// TIA Portal project "oscat_basic_332_s7_TIA_V12_V13_SP1_V14_V15.1" (V15.1) (continued)
VERSION : 1.1
// GEN_PW2 generates a time TH? followed by a time TL?.
// the input ts selects between 2 sets of timings for the operation.
// 
// uses: T_PLC_MS [FC64]
//       STIME [FB64],IDB_STIME [DB64]
   VAR_INPUT
      ENQ : Bool;
      TH1 : Time;
      TL1 : Time;
      TH2 : Time;
      TL2 : Time;
      TS : Bool;
   END_VAR
   VAR_OUTPUT
      Q : Bool;
      TH : Time;
      TL : Time;
   END_VAR
   VAR
      t_high : Time;
      t_low : Time;
      tx : Time;
      start : Time;
      init : Bool;
      et : Time;
   END_VAR
BEGIN


   (* read system timer *)
   #tx := T_CONV(DWORD_TO_DINT("T_PLC_MS"()));

   (* startup initialization *)
   IF NOT #init THEN
       #start := #tx;
       #init := TRUE;
       #TH := T#0s;
       #TL := T#0s;
   END_IF;

   (* timing selection *)
   IF #TS THEN
       #t_high := #TH2;
       #t_low := #TL2;
   ELSE
       #t_high := #TH1;
       #t_low := #TL1;
   END_IF;

   (* normal operation *)
   IF #ENQ THEN
       #et := #tx - #start;
       IF NOT #Q THEN
           IF #et >= #t_low THEN
               #Q := TRUE;
               #start := #tx;
               #TL := T#0s;
           ELSE
               #TL := #et;
           END_IF;
       ELSE
           IF #et >= #t_high THEN
               #Q := FALSE;
               #start := #tx;
               #TH := T#0s;
           ELSE
               #TH := #et;
           END_IF;
       END_IF;
   ELSE
       #Q := FALSE;
       #TH := T#0s;
       #TL := T#0s;
       #start := #tx;
   END_IF;


   (* revision history
   hm  26. sep. 2008   rev 1.0
       original version

   hm  14. mar. 2009   rev 1.1
       removed double assignments

   *)
END_FUNCTION_BLOCK

FUNCTION_BLOCK "GEN_RDM"   // FB97, SCL
TITLE = GEN_RDM
{ S7_Optimized_Access := 'FALSE' }
AUTHOR : oscat
FAMILY : SIGGEN
NAME : GEN_RDM
VERSION : 1.1
// this signal generator generates a random output. The signal is defined by period time (PT), 
// amplitude (AM), offset (OS).
// The Output waveform will have its max peak at AM/2 + OS and its minimum peak at -AM/2 + OS. 
// The period time PT defines how often the output signal will jump to a new randow value.
// The Output Q will be true for one cycle anytime the output OUT has changed
// 
// uses: T_PLC_MS [FC64]
//       STIME [FB64],IDB_STIME [DB64]
//       RDM [FC101]
//       BIT_COUNT [FC291] 
//       FRACT [FC83]
   VAR_INPUT
      PT : Time;
      AM : Real := 1.0e+0;
      OS : Real;
   END_VAR
   VAR_OUTPUT
      Q : Bool;
      Out : Real;
   END_VAR
   VAR
      tx : Time;
      last : Time;
      init : Bool;
   END_VAR
BEGIN


     (* read system time and prepare input data *)
     #tx := T_CONV(DWORD_TO_DINT("T_PLC_MS"())) - #last;

     (* init section *)
     IF NOT #init THEN
       #init := TRUE;
       #last := #tx;
       #tx := t#0s;
     END_IF;

     (* add last if one cycle is finished *)
     IF #tx >= #PT THEN
       #last := #last + #PT;
       #tx := #tx - #PT;

       (* generate output signal *)
       #Out := #AM * ("RDM"(0.0) - 0.5) + #OS;
       #Q := TRUE;
     ELSE
       #Q := FALSE;
     END_IF;

   (* revision history

   hm  7.2.2007    rev 1.0
     original version

   hm  16.9.2007    rev 1.1
     changes time() to T_plc_ms() for compatibility reasons

   *)
END_FUNCTION_BLOCK

FUNCTION_BLOCK "GEN_RDT"   // FB98, SCL
TITLE = GEN_RDT
{ S7_Optimized_Access := 'FALSE' }
AUTHOR : Schohaus
FAMILY : SIGGEN
NAME : GEN_RDT
VERSION : 1.1
// RDMT generates a defined pulse with pulse width TP_Q at random times. the random time will be defined with an minimum and maximum time.
// 
// uses: RDM [FC101]
//       T_PLC_MS [FC64] 
//       STIME [FB64],IDB_STIME [DB64] 
//       BIT_COUNT [FC291] 
//       FRACT [FC83]
   VAR_INPUT
      Enable : Bool := TRUE;
      Min_Time_ms : Time := T#1S;
      Max_Time_ms : Time := T#1S200MS;
      TP_Q : Time := T#100MS;
   END_VAR
   VAR_OUTPUT
      xQ : Bool;
   END_VAR
   VAR
      tonRDMTimer : TON;
      tof_xQ : TOF;
      tRDMTime : Time;
      rRDMTime : Real;
   END_VAR
BEGIN


   (*
   FUNCTION_BLOCK RDMTimer
   ###############################################################################
        Ersteller / author :                    J.Schohaus
        Datum / date:                         13.07.2007
   ###############################################################################
        Änderungen / Datum / Ersteller :                                                            
        moditication / date / author :        
   ###############################################################################
        Verwendete Bibliotheken     ( * werden im Baustein nicht benötigt )
                    Oscat.lib
   ###############################################################################
   Beschreibung:
   *)

     #tonRDMTimer ( IN:= #Enable , PT:= #tRDMTime );
     #tof_xQ ( IN:= #tonRDMTimer.Q , PT:= #TP_Q );
     #xQ := #tof_xQ.Q;
     IF #tonRDMTimer.Q THEN
          #xQ := TRUE ;
          #rRDMTime := "RDM" ( last:= #rRDMTime ) ;
          #tRDMTime := T_CONV(REAL_TO_DINT(#rRDMTime * DINT_TO_REAL(T_CONV(#Max_Time_ms - #Min_Time_ms)) + DINT_TO_REAL(T_CONV(#Min_Time_ms )))) ;
          #tonRDMTimer. IN:= FALSE ;
     END_IF;

   (* revision history
   J. Schohaus 19. nov 2007    rev 1.0
       origial version

   hm  16. mar. 2008           rev 1.1
       added type conversion to avoid warnings under codesys 3.0
   *)
END_FUNCTION_BLOCK

FUNCTION_BLOCK "GEN_RMP"   // FB99, SCL
TITLE = GEN_RMP
{ S7_Optimized_Access := 'FALSE' }
AUTHOR : oscat
FAMILY : SIGGEN
NAME : GEN_RMP
VERSION : 1.4
// this signal generator generates a ramp wave output. The ramp wave signal is defined by period time (PT), 
// amplitude (AM), offset (OS) and a specific delay for the output signal (DL).
// The Output waveform will have its minimum peak at OS and its maximum peak at AM + OS. 
// The delay input can delay a signal up to PT, this can be useful to synchronize different generators 
// and generate interleaving signals.
// in addition to the analog output Out there is a second boolean output Q with is true for one cycle when the ramp starts.
// 
// uses: T_PLC_MS [FC64]
//       STIME [FB64],IDB_STIME [DB64]
//       MODR [FC97]
//       FLOOR2 [FC82] 
//       FRACT [FC83]
//       MULTIME [FC203]
   VAR_INPUT
      PT : Time := T#1S;
      AM : Real := 1.0e+0;
      OS : Real;
      DL : Real;
   END_VAR
   VAR_OUTPUT
      Q : Bool;
      OUT : Real;
   END_VAR
   VAR
      tx : Time;
      last : Time;
      init : Bool;
      temp : Real;
      ltemp : Real;
   END_VAR
BEGIN


   (* read system time and prepare input data *)
   #tx := T_CONV(DWORD_TO_DINT("T_PLC_MS"())) - #last;
   #DL := "MODR"(IN:=#DL,DIVI:=1.0);
   IF #DL < 0.0 THEN #DL := 1.0 - #DL; END_IF;

   (* init section *)
   IF NOT #init THEN
       #init := TRUE;
       #last := #tx;
       #tx := t#0s;
   END_IF;

   (* add last if one cycle is finished *)
   IF #tx >= #PT THEN
       #last := #last + #PT;
       #tx := #tx - #PT;
   END_IF;

   (* generate sine wave *)
   #ltemp := #temp;
   IF #PT > t#0s THEN #temp := "FRACT"(DINT_TO_REAL(T_CONV(#tx + "MULTIME"(t:=#PT,M:=#DL))) / DINT_TO_REAL(T_CONV(#PT))); END_IF;
   #OUT := #AM * #temp + #OS;

   (* boolean output Q *)
   #Q := #temp < #ltemp;


   (* revision history
   hm  3. mar 2007     rev 1.0
       original version

   hm  17 sep 2007     rev 1.1
       replaced time() with t_plc_ms for compatibilitx reasons

   hm  27. nov 2007    rev 1.2
       avoid divide by 0 when pt = 0

   ks  26. oct. 2008   rev 1.3
       code optimization

   hm  10. mar. 2009   rev 1.4
       changed real constants to use dot syntax
   *)
END_FUNCTION_BLOCK

FUNCTION_BLOCK "GEN_SIN"   // FB100, SCL
TITLE = GEN_SIN
{ S7_Optimized_Access := 'FALSE' }
AUTHOR : oscat
FAMILY : SIGGEN
NAME : GEN_SIN
VERSION : 1.6
// this signal generator generates a sine wave output. The sine wave signal is defined by period time (PT), 
// amplitude (AM), offset (OS) and a specific delay for the output signal (DL).
// The Output waveform will have its max peak at AM/2 + OS and its minimum peak at -AM/2 + OS. 
// The delay input can delay a signal up to PT, this can be useful to synchronize different generators 
// and generate interleaving signals. A Cos wave can be generated accordingly.
// in addition to a analog output Out there is a second boolean output Q with the corresponding binary signal.
//  
// uses: T_PLC_MS [FC64]
//       STIME [FB64],IDB_STIME [DB64]
//       MODR [FC97]
//       FLOOR2 [FC82] 
//       MULTIME [FC203]
//       SIGN_R [FC109]
   VAR_INPUT
      PT : Time;
      AM : Real := 1.0e+0;
      OS : Real;
      DL : Real;
   END_VAR
   VAR_OUTPUT
      Q : Bool;
      OUT : Real;
   END_VAR
   VAR
      tx : Time;
      last : Time;
      init : Bool;
      temp : Real;
   END_VAR
BEGIN


   (* read system time and prepare input data *)
   #tx := T_CONV(DWORD_TO_DINT("T_PLC_MS"())) - #last;
   #DL := "MODR"(IN:=#DL,DIVI:=1.0);
   IF #DL < 0.0 THEN #DL := 1.0 - #DL; END_IF;

   (* init section *)
   IF NOT #init THEN
       #init := TRUE;
       #last := #tx;
       #tx := t#0s;
   END_IF;

   (* add last if one cycle is finished *)
   IF #tx >= #PT THEN
       #last := #last + #PT;
       #tx := #tx - #PT;
   END_IF;

   (* generate sine wave *)
   IF #PT > t#0s THEN #temp := SIN("PI2" * DINT_TO_REAL(T_CONV(#tx + "MULTIME"(t:=#PT,M:=#DL))) / DINT_TO_REAL(T_CONV(#PT))); END_IF;
   #OUT := #AM * 0.5 *  #temp + #OS;

   (* boolean output Q *)
   #Q := NOT "SIGN_R"(#temp);


   (* revision history
   hm  22. jan 2007    rev 1.0
       original version

   hm  17 sep 2007 rev 1.1
       replaced time() with t_plc_ms for compatibilitx reasons

   hm  27. nov 2007    rev 1.2
       avoid divide by 0 when pt = 0

   hm  6. jan 2008     rev 1.3
       improved performance

   hm  16. mar. 2008   rev 1.4
       added type conversion to avoid warnings under codesys 3.0

   hm  18. oct. 2008   rev 1.5
       using math constants

   hm  11. mar. 2009   rev 1.6
       changed real constants to use dot syntax

   *)
END_FUNCTION_BLOCK

FUNCTION_BLOCK "GEN_SQR"   // FB101, SCL
TITLE = GEN_SQR
{ S7_Optimized_Access := 'FALSE' }
AUTHOR : oscat
FAMILY : SIGGEN
NAME : GEN_SQR
VERSION : 1.4
// this signal generator generates a square wave output. The square wave signal is defined by period time (PT), 
// amplitude (AM), offset (OS), duty cycle (DC) and a specific delay for the output signal (DL).
// The Output waveform will switch between AM/2 + OS and -AM/2 + OS. The DC input specifies ther duty cycle, 
// DC = 0 means output is low at all times and 1 means output is high at all times.
// The delay input can delay a signal up to PT, this can be useful to synchronize different generators and generate interleaving signals.
// in addition to a analog output Out there is a second boolean output Q.
// 
// uses: T_PLC_MS [FC64]
//       STIME [FB64],IDB_STIME [DB64]
//       MODR [FC97]
//       FLOOR2 [FC82] 
//       MULTIME [FC203]
   VAR_INPUT
      PT : Time;
      AM : Real := 1.0e+0;
      OS : Real;
      DC : Real := 5.0e-1;
      DL : Real;
   END_VAR
   VAR_OUTPUT
      Q : Bool;
      Out : Real;
   END_VAR
   VAR
      tx : Time;
      last : Time;
      init : Bool;
   END_VAR
BEGIN


   (* check dc = 1 or 0 *)
   IF #DC = 0.0 THEN
       #Out := -#AM * 0.5 + #OS;
       #Q := FALSE;
       RETURN;
   ELSIF #DC = 1.0 THEN
       #Out := #AM * 0.5 + #OS;
       #Q := TRUE;
       RETURN;
   END_IF;

   (* read system time and prepare input data *)
   #tx := T_CONV(DWORD_TO_DINT("T_PLC_MS"())) - #last;
   #DL := "MODR"(IN:=#DL,DIVI:=1.0);
   IF #DL < 0.0 THEN #DL := 1.0 - #DL; END_IF;
   #DC := "MODR"(IN:=#DC,DIVI:=1.0);
   IF #DC < 0.0 THEN #DC := 1.0 - #DC; END_IF;

   (* init section *)
   IF NOT #init THEN
       #init := TRUE;
       #last := #tx;
       #tx := t#0s;
   END_IF;

   (* add last if one cycle is finished *)
   IF #tx >= #PT THEN
       #last := #last + #PT;
       #tx := #tx - #PT;
   END_IF;

   (* check if falling or rising edge first *)
   IF "MULTIME"(t:=#PT,M:=#DL + #DC) >= #PT THEN
       (* generate falling edge *)
       IF #tx >= "MULTIME"(t:=#PT,M:=#DL + #DC - 1) THEN
           #Out := -#AM * 0.5 + #OS;
           #Q := FALSE;
       END_IF;
       (* generate rising edge *)
       IF #tx >= "MULTIME"(t:=#PT,M:=#DL) THEN
           #Out := #AM * 0.5 + #OS;
           #Q := TRUE;
       END_IF;
   ELSE
       (* generate rising edge first *)
       IF #tx >= "MULTIME"(t:=#PT,M:=#DL) THEN
           #Out := #AM * 0.5 + #OS;
           #Q := TRUE;
       END_IF;
       (* generate falling edge *)
       IF #tx >= "MULTIME"(t:=#PT,M:=#DL + #DC) THEN
           #Out := -#AM * 0.5 + #OS;
           #Q := FALSE;
       END_IF;
   END_IF;


   (* revision history

   hm  12. feb 2007    rev 1.1
       added default value for dc = 0.5

   hm  17 sep 2007 rev 1.2
       replaced time() with t_plc_ms for compatibilitx reasons

   hm  6. jan 2008 rev 1.3
       improved performance

   hm  11. mar. 2009   rev 1.4
       changed real constants to use dot syntax
       set default amplitude to 1.0

   *)
END_FUNCTION_BLOCK

FUNCTION_BLOCK "PWM_DC"   // FB102, SCL
TITLE = PWM_DC
{ S7_Optimized_Access := 'FALSE' }
AUTHOR : oscat
FAMILY : SIGGEN
NAME : PWM_DC
VERSION : 1.4
// this signal generator generates a square wave signal which is specified by the frequency and the duty cycle
// 
// uses: CLK_PRG [FB52]
//       T_PLC_MS [FC64] 
//       STIME [FB64],IDB_STIME [DB64] 
//       TP_X [FB69]
   VAR_INPUT
      F : Real;
      DC : Real;
   END_VAR
   VAR_OUTPUT
      Q : Bool;
   END_VAR
   VAR
      clk : "CLK_PRG";
      pulse : "TP_X";
   END_VAR
   VAR_TEMP
      tmp : Real;
   END_VAR
BEGIN


   IF #F > 0.0 THEN
       #tmp := 1000.0 / #F;
       #clk(PT := T_CONV(REAL_TO_DINT(#tmp)));
       #pulse(IN := #clk.Q, PT := T_CONV(REAL_TO_DINT(#tmp * #DC)));
       #Q := #pulse.Q;
   END_IF;


   (* revision history

   hm  25. feb 2007    rev 1.1
       recoded in st for better performance and better portability

   hm  27. nov 2007    rev 1.2
       avoid divide by 0 when F = 0

   hm  19. oct. 2008   rev 1.3
       changed type TP_R to TP_X because of name change
       improved performance

   hm  11. mar. 2009   rev 1.4
       changed real constants to use dot syntax

   *)
END_FUNCTION_BLOCK

FUNCTION_BLOCK "PWM_PW"   // FB103, SCL
TITLE = PWM_PW
{ S7_Optimized_Access := 'FALSE' }
AUTHOR : oscat
FAMILY : SIGGEN
NAME : PWM_PW
VERSION : 1.5
// this signal generator generates a square wave signal which is specified by the frequency and the pulse width.
// 
// uses: CLK_PRG [FB52]
//       T_PLC_MS [FC64] 
//       STIME [FB64],IDB_STIME [DB64] 
//       TP_X [FB69]
   VAR_INPUT
      F : Real;
      PW : Time;
   END_VAR
   VAR_OUTPUT
      Q : Bool;
   END_VAR
   VAR
      clk : "CLK_PRG";
      pulse : "TP_X";
   END_VAR
BEGIN


   IF #F > 0.0 THEN
       #clk(PT := T_CONV(REAL_TO_DINT(1000.0 / #F)));
       #pulse(IN := #clk.Q, PT := #PW);
       #Q := #pulse.Q;
   END_IF;


   (* revision history

   hm  25. feb 2007    rev 1.1
       recoded in st for better performance and better portability

   hm  27. nov 2007    rev 1.2
       avoid divide by 0 when F = 0

   hm  9. dec 2007     rev 1.3
       corrected an error with F = 0

   hm  19. oct. 2008   rev 1.4
       changed type tp_r to TP_x brecause of name change

   hm  11. mar. 2009   rev 1.5
       changed real constants to use dot syntax

   *)
END_FUNCTION_BLOCK

FUNCTION_BLOCK "RMP_SOFT"   // FB104, SCL
TITLE = RMP_SOFT
{ S7_Optimized_Access := 'FALSE' }
AUTHOR : oscat
FAMILY : SIGGEN
NAME : RMP_SOFT
VERSION : 2.0
// this soft on/off ramp generator generates a soft on and soft off ramp while the max on value is set by the input
// the time for a full ramp can be set by config variables for up and down ramp.
// 
// uses: _RMP_B [FB93]
//       T_PLC_MS [FC64] 
//       STIME [FB64],IDB_STIME [DB64]
   VAR_INPUT
      IN : Bool;
      VAL : Byte;
      PT_ON : Time;
      PT_OFF : Time;
   END_VAR
   VAR_OUTPUT
      OUT : Byte;
   END_VAR
   VAR
      rmp : "_RMP_B";
      tmp : Byte;
   END_VAR
BEGIN


   #tmp := INT_TO_BYTE(SEL(G:=#IN, IN0:=0, IN1:=BYTE_TO_INT(#VAL)));
   IF BYTE_TO_INT(#tmp) > BYTE_TO_INT(#OUT) THEN
       (* we need to ramp down *)
       #rmp(DIR := TRUE, E := TRUE, TR := #PT_ON, RMP := #OUT);
       (* make sure out does not surpass tmp *)
       #OUT := INT_TO_BYTE(MIN(IN1:=BYTE_TO_INT(#OUT), IN2:=BYTE_TO_INT(#tmp)));
   ELSIF BYTE_TO_INT(#tmp) < BYTE_TO_INT(#OUT) THEN
       (* we need to ramp up *)
       #rmp(DIR := FALSE, E := TRUE, TR := #PT_OFF, RMP := #OUT);
       (* make sure out does not surpass tmp *)
       #OUT := INT_TO_BYTE(MAX(IN1:=BYTE_TO_INT(#OUT), IN2:=BYTE_TO_INT(#tmp)));
   ELSE
       (* no ramp necessary *)
       #rmp(E := FALSE, RMP := #OUT);
   END_IF;


   (* revision history

   hm 22.1.2007    rev 1.1
       deleted unused variables X1 and I, X2 and X3

   hm  17.9.2007   rev 1.2
       replaced time() with t_plc_ms() for compatibility reasons

   hm  26. oct. 2008   2.0
       new code using _rmp_b
   *)
END_FUNCTION_BLOCK

FUNCTION_BLOCK "RMP_W"   // FB105, SCL
TITLE = RMP_W
{ S7_Optimized_Access := 'FALSE' }
AUTHOR : oscat
FAMILY : SIGGEN
NAME : RMP_W
VERSION : 2.0
// this ramp generator generates a Word wide ramp with 65535 steps
// the generator has an asynchronous set and reset
// the ramp is controlled by PT which is the total ramp time for a full sweep from 0..65535
// an UD input controlls the direction Up or Down and the E input enables the ramp generation
// a busy output indicates that the ramp is running, busy false means output is stable.
// the outputs low and high will be true when the output has reached its max or min value.
// 
// uses: _RMP_W [FB94]
//       T_PLC_MS [FC64] 
//       STIME [FB64],IDB_STIME [DB64]
   VAR_INPUT
      SET : Bool;
      PT : Time;
      "E" : Bool := TRUE;
      UP : Bool := TRUE;
      RST : Bool;
   END_VAR
   VAR_OUTPUT
      out : Word;
      busy : Bool;
      high : Bool;
      low : Bool;
   END_VAR
   VAR
      rmp : "_RMP_W";
   END_VAR
BEGIN


   #rmp(DIR := #UP, E := #"E", TR := #PT, RMP := #out);

   (* set or reset operation *)
   IF #RST THEN
       #out := 0;
   ELSIF #SET THEN
       #out := 65535;
   END_IF;

   (* checks for outputs stable and reset or set busy flag *)
   #low := #out = 0;
   #high := #out = 65535;
   #busy := NOT (#low OR #high) AND #"E";


   (* revision history:

   hm 4.10.2006        rev 1.1
       added the busy output which signals that the ramp is running.

   hm 22.1.2007        rev 1.2
       deleted unused variable step

   hm  17.9.2007       rev 1.3
       replaced time() with t_plc_ms() for compatibility reasons

   hm  28. sep 2007    rev 1.4
       added outputs on and off
       busy is now disabled while en is false
       new coding for higher accuracy and performance

   hm  5. oct 2007 rev 1.5
       added statements to allow for PT to be t#0s output jumps to max or min immediately

   hm  2. dec 2007 rev 1.6
       corrected an error in calculation of step response

   hm  25. dec 2007    rev 1.7
       corrected an error while step response was too slow for fast rise times

   hm  16. oct. 2008   rev 1.8
       improved performance

   hm  18. oct. 2008   rev 1.9
       renamed inout EN to E for compatibility reasons

   hm  23. oct. 2008   rev 2.0
       new code using _RMP_W
   *)
END_FUNCTION_BLOCK

FUNCTION_BLOCK "RMP_B"   // FB232, SCL
TITLE = RMP_B
{ S7_Optimized_Access := 'FALSE' }
AUTHOR : oscat
FAMILY : SIGGEN
NAME : RMP_B
VERSION : 2.0
// this ramp generator generates a byte wide ramp with 255 steps
// the generator has an asynchronous set and reset
// the ramp is controlled by PT which is the total ramp time for a full sweep from 0..255
// an UD input controlls the direction Up or Down and the E input enables the ramp generation
// a busy output indicates that the ramp is running, busy false means output is stable.
// the outputs low and high will be true when the output has reached its max or min value.
// 
// uses: _RMP_B [FB93]
//       T_PLC_MS [FC64] 
//       STIME [FB64],IDB_STIME [DB64]
   VAR_INPUT
      SET : Bool;
      PT : Time;
      "E" : Bool := TRUE;
      UP : Bool := TRUE;
      RST : Bool;
   END_VAR
   VAR_OUTPUT
      OUT : Byte;
      BUSY : Bool;
      HIGH : Bool;
      LOW : Bool;
   END_VAR
   VAR
      rmp : "_RMP_B";
   END_VAR
BEGIN


   (* generate ramp *)
   #rmp(DIR := #UP, E := #"E", TR := #PT, RMP := #OUT);

   (* set or reset operation *)
   IF #RST THEN
       #OUT := 0;
   ELSIF #SET THEN
       #OUT := 255;
   END_IF;

   (* checks for outputs stable and reset or set busy flag *)
   #LOW := #OUT = 0;
   #HIGH := #OUT = 255;
   #BUSY := NOT (#LOW OR #HIGH) AND #"E";


   (* revision history

   hm 5.10.2006    rev 1.1
       added busy output
   hm 17.1.2007    rev 1.2
       renamed input ud to up for better usability
       deleted unused variable step

   hm  17.9.2007       rev 1.3
       replaced time() with t_plc_ms() for compatibility reasons

   hm  28. sep 2007    rev 1.4
       added outputs on and off
       busy is now disabled while en is false
       new coding for higher accuracy and performance

   hm  5. oct 2007 rev 1.5
       added statements to allow for PT to be t#0s output jumps to max or min immediately

   hm  25. dec 2007    rev 1.6
       improved code for better performance

   hm  16. oct. 2008   rev 1.7
       improved code for better performance

   hm  18. oct. 2008   rev 1.8
       added type conversion to avoid warnings
       changed input en to e for compatibility reasons

   hm  23. oct. 2008   REV     2.0
       new code using _RMP_B

   *)
END_FUNCTION_BLOCK

FUNCTION_BLOCK "TREND_DW"   // FB245, SCL
TITLE = TREND_DW
{ S7_Optimized_Access := 'FALSE' }
AUTHOR : hugo
FAMILY : SIGPRO
NAME : TREND_DW
VERSION : 1.2
// trend_DW analyses the trend of a input signal.
// The Output Q is True if the input X is >= last_X and is false if the input X is <= last_X
// in addition to the trend the output TU will be high for one cycle to signal a rising of the input value X
// and  TD will signal a decreasing value on the input X.
// in case of a change the output D will show the delta of the input to the last input value.
   VAR_INPUT
      X : DWord;
   END_VAR
   VAR_OUTPUT
      Q : Bool;
      TU : Bool;
      TD : Bool;
      D : DWord;
   END_VAR
   VAR
      last_X : DWord;
   END_VAR
BEGIN


   IF DWORD_TO_DINT(#X) > DWORD_TO_DINT(#last_X) THEN
       #TU := TRUE;
       #TD := FALSE;
       #D := DINT_TO_DWORD(DWORD_TO_DINT(#X) - DWORD_TO_DINT(#last_X));
       #Q := TRUE;
   ELSIF DWORD_TO_DINT(#X) < DWORD_TO_DINT(#last_X) THEN
       #TD := TRUE;
       #TU := FALSE;
       #D := DINT_TO_DWORD(DWORD_TO_DINT(#last_X) - DWORD_TO_DINT(#X));
       #Q := FALSE;
   ELSE
       #TU := FALSE; 
       #TD := FALSE;
       #D := 0;
   END_IF;
   #last_X := #X;


   (* revision history
   hm  21. nov. 2008   rev 1.0
       original version

   hm  20. feb. 2009   rev 1.1
       added outputs TU, TD and D

   hm  14. mar. 2009   rev 1.2
       removed double assignments

   *)
END_FUNCTION_BLOCK

FUNCTION_BLOCK "_RMP_NEXT"   // FB246, SCL
TITLE = _RMP_NEXT
{ S7_Optimized_Access := 'FALSE' }
AUTHOR : hugo
FAMILY : SIGGEN
NAME : RMP_NEXT
VERSION : 1.4
// _RMP_NEXT  will generate a ramp output following the input IN.
// on a rising ramp the output will stop as soon as it has surpassed the input in, and on a falling ramp it will stop when out is smaller than in.
// a lockout time T_L will be added between up and down direction.
// 
// uses: _RMP_B [FB93]
//       TREND_DW [FB245]
//       T_PLC_MS [FC64]
//       STIME [FB64],IDB_STIME [DB64]
   VAR_INPUT
      "E" : Bool := TRUE;
      IN : Byte;
      TR : Time;
      TF : Time;
      TL : Time;
   END_VAR
   VAR_OUTPUT
      DIR : Bool;
      UP : Bool;
      DN : Bool;
   END_VAR
   VAR_IN_OUT
      OUT : Byte;
   END_VAR
   VAR
      rmx : "_RMP_B";
      dirx : "TREND_DW";
      t_lock : TP;
      xen : Bool;
      xdir : Bool;
   END_VAR
BEGIN


   #dirx(X := #IN);

   #t_lock(IN := FALSE, PT := #TL);

   IF #dirx.TU AND (BYTE_TO_INT(#OUT) < BYTE_TO_INT(#IN)) THEN
       IF NOT #xdir AND #xen THEN #t_lock.IN := TRUE; END_IF;
       #xen := TRUE;
       #xdir := TRUE;
   ELSIF #dirx.TD AND (BYTE_TO_INT(#OUT) > BYTE_TO_INT(#IN)) THEN
       IF #xdir AND #xen THEN #t_lock.IN := TRUE; END_IF;
       #xen := TRUE;
       #xdir := FALSE;
   ELSIF #xen THEN
       IF (#xdir AND (BYTE_TO_INT(#OUT) >= BYTE_TO_INT(#IN))) OR (NOT #xdir AND (BYTE_TO_INT(#OUT) <= BYTE_TO_INT(#IN))) THEN
           #xen := FALSE;
           IF #TL > t#0s THEN #t_lock.IN := TRUE; END_IF;
       END_IF;
   END_IF;

   IF NOT #t_lock.Q AND #xen THEN
       #UP := #xdir; 
       #DIR := #xdir;
       #DN := NOT #xdir;
   ELSE
       #DN := FALSE;
       #UP := FALSE; 
   END_IF;

   #rmx(RMP := #OUT, E := #"E" AND (#UP OR #DN) , DIR := #DIR, TR := SEL(G:=#DIR, IN0:=#TF, IN1:=#TR));


   (* revison history
   hm  23. nov. 2008 rev 1.0
     original version

   hm  24. jan. 2009 rev 1.1
     deleted unused vars tmp1, tmp2

   hm  20. feb. 2009 rev 1.2
     improved algorithm
     added TL

   hm  9. mar. 2009  rev 1.3
     input E was ignored
     removed double assignments

   hm  18. jul. 2009 rev 1.4
     improved performance

   *)
END_FUNCTION_BLOCK

FUNCTION "T_PLC_MS" : DWord   // FC64, SCL
TITLE = T_PLC_MS
{ S7_Optimized_Access := 'FALSE' }
AUTHOR : hugo
FAMILY : MEASURE
NAME : T_PLC_MS
VERSION : 1.2
// T_PLC_MS reads the internal PLC timer and return the time, it has the advantage to be able to set a debug mode 
// and speed up the counter to test the plc timer overrun which occurs every 50 days respectively 25 days at siemens S7
// this routine also allows to correct the behavior of s7 where the internal plc counter will not count all 32 bits.
// 
// uses: STIME [FB64],IDB_STIME [DB64]
BEGIN


   "IDB_STIME"(); 
   #T_PLC_MS := "IDB_STIME".tx; 
   (* hier muss die korrektur für step7 stattfinden
   plctime muss den vollen wertebereich von time ausnutzen:
   wenn bei step7 time -24tage bis plus 24 tage ist dann muss der timer auch beim überlauf auf -24tage springen 
   und auf keinen fall auf 0 !!!!
   für siemens muss ein weiterer fb im main eingebunden werden der sicherstellt das alle 32 bits durchgezählt werden.
   es kann nur ein fb sein den er muss sich das oberste (32te) bit merken.
   oder etwa spring s7 bei überlauf auf -24 tage????? dann wäre keine korrektur nötig.
   *)
   IF "debug" THEN
       #T_PLC_MS := DINT_TO_DWORD((DWORD_TO_DINT(SHL(IN:=#T_PLC_MS,N:="N") OR SHL(IN:=DWORD#1,N:="N"))-1) + DWORD_TO_DINT("offset_1"));
   END_IF;


   (* revision history
   hm  14.9.2007   rev 1.0
       original version

   hm  12. nov 2007    rev 1.1
       added temporaray variable tx because some compilers could not handle time() as an argument

   hm  16. nov. 2008   rev 1.2
       initialized constants with 0 for compatibility reasons
   *)
END_FUNCTION

FUNCTION "FLOOR2" : DInt   // FC82, SCL
TITLE = FLOOR2
{ S7_Optimized_Access := 'FALSE' }
AUTHOR : hugo
FAMILY : MATH
NAME : FLOOR2
VERSION : 1.1
// This is a rounding function which returns the biggest possible integer which is less or equal to X.
// floor2(3.14) = 3
// floor2(-3.14) = -4
   VAR_INPUT
      X : Real;
   END_VAR
BEGIN


   #FLOOR2 := REAL_TO_DINT(#X);
   IF DINT_TO_REAL(#FLOOR2) > #X THEN
     #FLOOR2 := #FLOOR2 - 1;
   END_IF;

   (* revision history
   hm  21. mar. 2008   rev 1.0
       originlal version

   hm  4. apr. 2008    rev 1.1
       added type conversion to avoid warnings under codesys 3.0
   *)
END_FUNCTION

FUNCTION "FRACT" : Real   // FC83, SCL
TITLE = FRACT
{ S7_Optimized_Access := 'FALSE' }
AUTHOR : hugo
FAMILY : MATH
NAME : FRACT
VERSION : 1.3
// this function returns the fraction of a real number
// fract(3.14) = 0.14
   VAR_INPUT
      x : Real;
   END_VAR
BEGIN


   IF ABS(#x) < 2.0E9 THEN
       #FRACT := #x - DINT_TO_REAL(TRUNC(#x));
   ELSE
       #FRACT := 0.0;
   END_IF;


   (* revision history
   hm  4. aug 2006 rev 1.0
       original version

   hm  11. mar 2008    rev 1.1
       added dint_to_real for compatibility reasons
       now returns 0 for number > 2e9
       changed input to x

   hm  21. mar. 2008   rev 1.2
       use D_trunc instead of TRUNC for compatibility reasons

   hm  10. mar. 2009   rev 1.3
       real constants updated to new systax using dot

   *)
END_FUNCTION

FUNCTION "MODR" : Real   // FC97, SCL
TITLE = MODR
{ S7_Optimized_Access := 'FALSE' }
AUTHOR : hugo
FAMILY : MATH
NAME : MODR
VERSION : 1.5
// this is a modulo funtion for real numbers
// modr(5.5,2.5) = 0.5
// 
// uses: FLOOR2 [FC82]
   VAR_INPUT
      IN : Real;
      DIVI : Real;
   END_VAR
BEGIN


   IF #DIVI = 0.0 THEN
       #MODR := 0.0;
   ELSE
       #MODR := #IN - DINT_TO_REAL("FLOOR2"(#IN / #DIVI)) * #DIVI;
   END_IF;


   (* revision history

   hm  4. aug.2006     rev 1.0

   hm  28. jan.2007   rev 1.1
       modr(x,0) will deliver the result 0

   hm  21. mar 2008    rev 1.2
       use D_trunc for compatibility reasons

   hm  4. apr. 2008    rev 1.3
       added type conversion to avoid warnings under codesys 3.0

   hm  31. oct. 2008   rev 1.4
       changed algorithm to the more common version using floor instead of TRUNC

   hm  10. mar. 2009   rev 1.5
       real constants updated to new systax using dot

   *)
END_FUNCTION

FUNCTION "RDM" : Real   // FC101, SCL
TITLE = RDM
{ S7_Optimized_Access := 'FALSE' }
AUTHOR : hugo
FAMILY : MATH
NAME : RDM
VERSION : 1.9
// this function calculates a pseudo random number
// to generate the number it reads the sps timer and calculates a random number between 0 and 1:
// in order to use rdm more then once within one sps cycle it need to be called with different seed numbers LAST.
//  
// uses: T_PLC_MS [FC64]
//       STIME [FB64],IDB_STIME [DB64]
//       BIT_COUNT [FC291]
//       FRACT [FC83]
   VAR_INPUT
      last : Real;
   END_VAR
   VAR_TEMP
      tn : DWord;
      _tn AT tn : Array[0..31] of Bool;
      tc : Int;
   END_VAR
BEGIN


   #tn := "T_PLC_MS"();
   #tc := "BIT_COUNT"(#tn);
   #_tn[7] := #_tn[26];  //tn.31 := tn.2;
   #_tn[6] := #_tn[29];  //tn.30 := tn.5;
   #_tn[5] := #_tn[28];  //tn.29 := tn.4;
   #_tn[4] := #_tn[25];  //tn.28 := tn.1;
   #_tn[3] := #_tn[24];  //tn.27 := tn.0;
   #_tn[2] := #_tn[31];  //tn.26 := tn.7;
   #_tn[1] := #_tn[30];  //tn.25 := tn.6;
   #_tn[0] := #_tn[27];  //tn.24 := tn.3;
   #tn := ROL(IN:=#tn,N:="BIT_COUNT"(#tn)) AND 16#7FFFFFFF OR 16#40000001;  // OR 16#80000001
   #tn := DINT_TO_DWORD(DWORD_TO_DINT(#tn) MOD 71474513 + #tc + 77);
   #RDM := "FRACT"(DINT_TO_REAL(DWORD_TO_DINT(#tn)) / 10000000.0 * ("E"- LIMIT(MN:=0.0,IN:=#last,MX:=1.0)));


   (*
   pt := ADR(temp);
   pt^ := (T_PLC_MS() AND 16#007FFFFF) OR 16#3D000000;
   RDM := fract(modR(temp*e+pi1, PI1-last) + modR(temp*PI1+e + last,e-last));
   *)

   (* revision history
   hm      16. jan 2007        rev 1.0
       original version

   hm      11. nov 2007        rev 1.1
       changed time() into t_plc_ms()

   hm      20. nov 2007        rev 1.2
       changed code of temp calculation to avoid overflow in modr due to resuclt would not fit DINT for high timeer values

   hm      5. jan 2008     rev 1.3
       changed calculation of temp to avoid problem with high values of t_plc_ms

   hm      2. feb 2008     rev 1.4
       changed algorithm to avoind non iec functions and guarantee more randomness

   hm  10. mar. 2008       rev 1.5
       make sure last will be between 0 and 1 to avoid invalid results

   hm  16. mar. 2008       rev 1.6
       added conversion for tc to avoid warnings under codesys 3.0

   hm  18. may. 2008       rev 1.7
       changed constant E to E1

   hm  18. oct. 2008       rev 1.8
       using math constants

   hm  10. mar. 2009       rev 1.9
       real constants updated to new systax using dot

   *)
END_FUNCTION

FUNCTION "SIGN_R" : Bool   // FC109, SCL
TITLE = SIGN_R
{ S7_Optimized_Access := 'FALSE' }
AUTHOR : hugo
FAMILY : MATH
NAME : SIGN_R
VERSION : 1.4
// this function return true if the real input is negative
   VAR_INPUT
      in : Real;
   END_VAR
BEGIN


   #SIGN_R := #in < 0.0;


   (* revision history
   hm 19.1.2007    rev 1.1
       changed method of function for better compatibility to other systems

   hm  1.12.2007   rev 1.2
       changed code to improve performance

   hm  14. jun. 2008   rev 1.3
       improved performace

   hm 10. mar. 2009    rev 1.4
       real constants updated to new systax using dot
   *)
END_FUNCTION

FUNCTION "MULTIME" : Time   // FC203, SCL
TITLE = MULTIME
{ S7_Optimized_Access := 'FALSE' }
AUTHOR : hugo
FAMILY : TIDT
NAME : MULTIME
VERSION : 1.1
// multiplies a time by a real number and returns a time
   VAR_INPUT
      t : Time;
      "M" : Real;
   END_VAR
BEGIN


     #MULTIME := T_CONV(REAL_TO_DINT(DINT_TO_REAL(T_CONV(#t))*#"M"));

   (* revision history
   hm      2. oct 2006 rev 1.0
       original version

   hm      14. mar 2008    rev 1.1
       rounded the result after the last digit

   *)
END_FUNCTION

FUNCTION "BIT_COUNT" : Int   // FC291, SCL
TITLE = BIT_COUNT
{ S7_Optimized_Access := 'FALSE' }
AUTHOR : hugo
FAMILY : GATE
NAME : BITCT
VERSION : 1.1
// BIT_COUNT counts the amount True of bits in a dword.
// for exabple: bit_count(3) returns 2 because two bits (bits 0 and 1) are true and all others are false.
   VAR_INPUT
      IN : DWord;
   END_VAR
   VAR_TEMP
      temp : DWord;
      attemp AT temp : Array[0..31] of Bool;
   END_VAR
BEGIN


     #BIT_COUNT := 0;
     #temp := #IN;

     WHILE DWORD_TO_DINT(#temp) <> 0 DO
       IF #attemp[24] THEN #BIT_COUNT := #BIT_COUNT +1; END_IF;
       #temp := SHR(IN:=#temp,N:=1);
     END_WHILE;

   (* revision history
   5.7.2007  rev 1.0    original version

   10.9.2007  rev 1.1    hm
     changed algorithm for better performace
     the execution time has reduced by a factor of 5
     deleted unused variable temp
   *)
END_FUNCTION

FUNCTION "FRMP_B" : Byte   // FC424, SCL
TITLE = FRMP_B
{ S7_Optimized_Access := 'FALSE' }
AUTHOR : hugo
FAMILY : FUNCT
NAME : FRMP_B
VERSION : 1.0
// this function calculates a ramp and limits the output to 0 .. 255 without overflow problems
   VAR_INPUT
      START : Byte;
      DIR : Bool;
      TD : Time;
      TR : Time;
   END_VAR
   VAR_TEMP
      tTD : Time;
   END_VAR
BEGIN


   #tTD := #TD;  // only Step7

   IF #TD < #TR THEN
     #FRMP_B := DINT_TO_BYTE(MIN(IN1:=DWORD_TO_DINT(SHL(IN:=DINT_TO_DWORD(T_CONV(#tTD)), N:=8)) / T_CONV(#TR) 
                                ,IN2:=SEL(G:=#DIR, IN0:=BYTE_TO_DINT(#START), IN1:=BYTE_TO_DINT(BYTE#255) - BYTE_TO_DINT(#START))));
     IF #DIR THEN
       #FRMP_B := INT_TO_BYTE(BYTE_TO_INT(#START) + BYTE_TO_INT(#FRMP_B));
     ELSE
       #FRMP_B := INT_TO_BYTE(BYTE_TO_INT(#START) - BYTE_TO_INT(#FRMP_B));
     END_IF;
   ELSE
     #FRMP_B := INT_TO_BYTE(DINT_TO_INT(SEL(G:=#DIR, IN0:=0, IN1:=255)));
   END_IF;


   (* revision history

   17. feb. 2011 rev 1.0
     new module

   *)
END_FUNCTION

// ===== PLC "Eng signal processing"  Unspecific CPU S7 300 =====

VAR_GLOBAL CONSTANT   // PLC tag table "STEP7 classic symbols"
   "debug" : Bool := FALSE;
   "N" : Int := 0;
   "offset_FC64" : Int := 0;   // MigChange: offset
   "ff" : DWord := 16#FFFFFFFF;
   "ff_FC318" : Byte := 2#1;   // MigChange: ff
   "offset_FC64_1" : DWord := 0;
END_VAR

DATA_BLOCK "IDB_STIME"   // DB64
{ S7_Optimized_Access := 'FALSE' }
AUTHOR : dalbi
FAMILY : MEASURE
VERSION : 0.0
// stored: InstanceOfName STIME
"STIME"
BEGIN
END_DATA_BLOCK

FUNCTION_BLOCK "STIME"   // FB64, SCL
TITLE = STIME
{ S7_Optimized_Access := 'FALSE' }
AUTHOR : dalbi
FAMILY : MEASURE
NAME : STIME
VERSION : 1.5
// this function block makes sure that the timer of a siemens sps counts from 0 - 2^32-1.
   VAR_OUTPUT
      tx : DWord;
      at_tx AT tx : Array[0..31] of Bool;
   END_VAR
   VAR
      last_time : DWord;
      bit31 : Bool;
      init : Bool := TRUE;
   END_VAR
   VAR_TEMP
      TOP_SI : Struct
         EV_CLASS : Byte;
         EV_NUM : Byte;
         PRIORITY : Byte;
         NUM : Byte;
         TYP2_3 : Byte;
         TYP1 : Byte;
         ZI1 : Word;
         ZI2_3 : DWord;
      END_STRUCT;
      START_UP_SI : Struct
         EV_CLASS : Byte;
         EV_NUM : Byte;
         PRIORITY : Byte;
         NUM : Byte;
         TYP2_3 : Byte;
         TYP1 : Byte;
         ZI1 : Word;
         ZI2_3 : DWord;
      END_STRUCT;
      ERR : Int;
   END_VAR
BEGIN


   (* this FB is only necessary for siemens sps
   the siemens sps timer counts from 0 to 2^31-1 and starts at 0 sfter overrun.
   this means that the bit 31 (the highest bit ) will never be used and therefore
   a problem arises when t2 - t1 is checked.
   t2 - t1 is always valid also in an timer overrun situation where the time t1 is very high and t2 is very low.
   the result of the subtraction t2 - t1 however is still valid.
   this calculation does not work for soiemens because the highest bit is not used.

   this module stores the highest bit, changes the highest bit at every overrun occurence and stuffs ther highest bit in the output.
   the output is then used by t_plc_us and t_plc_ms.

   the correction needs and fb and not a function because the value of the highest bit has to be stored.

   do never use this function block in a codesys environment. the timer in codesys is correct and runs from 0 to 2^32-1
   *)

   (* read actual startup info *)
   (* OB1_SCAN_1  BYTE  -  B#16#01: Abschluss des Neustarts (Warmstarts)
                        -  B#16#02: Abschluss des Wiederanlaufs
                        -  B#16#03: Abschluss des freien Zyklus
                        -  B#16#04: Abschluss des Kaltstarts
                        -  B#16#05: Erster OB 1-Zyklus der neuen Master-CPU nach 
                                    Master-Reserve-Umschaltung und STOP des 
                                    bisherigen Masters *)

   #ERR := RD_SINFO (TOP_SI => #TOP_SI, START_UP_SI => #START_UP_SI);

   (* reset last_time on system startup *)
   IF #TOP_SI.EV_NUM = 1 OR #TOP_SI.EV_NUM = 2 OR #TOP_SI.EV_NUM = 4 OR NOT #init THEN 
       #last_time := 0;
       #bit31 := false;
       #init := true;
   END_IF;

   (* read the system timer *)
   #tx := DINT_TO_DWORD(T_CONV(TIME_TCK()));

   (* stuff the highest bit into the timer value *)
   #at_tx[7] := #bit31;

   (* check for overrun *)
   IF DWORD_TO_DINT(#tx) < DWORD_TO_DINT(#last_time) THEN
       (* an overrun has occured, change the value of the highest bit *)
       #bit31 := NOT #bit31;
   END_IF;

   (* stuff the highest bit into the timer value *)
   #at_tx[7] := #bit31;

   (* remember the last system time for the next overrun check *)
   #last_time := #tx;


   (* revision history
   DA  14.9.2007 rev 1.0
     original version

   DA  24.2.2008 rev 1.1
     added self reset on system startup

   DA   2.5.2008 rev 1.2
     correct a problem running under OB35

   DA  12.3.2009 rev 1.3
     correct a problem run on different CPUs

   DA  22.12.2009 rev 1.4
     correct a problem on startup

   DA  19.09.2011 rev 1.5
     correct a error in code 
   *)
END_FUNCTION_BLOCK

FUNCTION_BLOCK "_RMP_W"   // FB94, SCL
TITLE = _RMP_W
{ S7_Optimized_Access := 'FALSE' }
AUTHOR : hugo
FAMILY : SIGGEN
NAME : _RMP_W
VERSION : 1.1
// _RMP_B generates a ramp on an external var of type byte
// tr is the total ramp time, E is an enable and dir the direction of the ramp
// 
// uses: T_PLC_MS [FC64]
//       STIME [FB64],IDB_STIME [DB64]
   VAR_INPUT
      DIR : Bool;
      "E" : Bool := TRUE;
      TR : Time;
   END_VAR
   VAR_IN_OUT
      RMP : Word;
   END_VAR
   VAR
      tx : DWord;
      tl : DWord;
      "step" : DInt;
      init : Bool;
      last_dir : Bool;
   END_VAR
   VAR_TEMP
      TOP_SI : Struct
         EV_CLASS : Byte;
         EV_NUM : Byte;
         PRIORITY : Byte;
         NUM : Byte;
         TYP2_3 : Byte;
         TYP1 : Byte;
         ZI1 : Word;
         ZI2_3 : DWord;
      END_STRUCT;
      START_UP_SI : Struct
         EV_CLASS : Byte;
         EV_NUM : Byte;
         PRIORITY : Byte;
         NUM : Byte;
         TYP2_3 : Byte;
         TYP1 : Byte;
         ZI1 : Word;
         ZI2_3 : DWord;
      END_STRUCT;
      ERR : Int;
   END_VAR
BEGIN


   (* read actual startup info *)
   (* OB1_SCAN_1  BYTE  -  B#16#01: Abschluss des Neustarts (Warmstarts)
                        -  B#16#02: Abschluss des Wiederanlaufs
                        -  B#16#03: Abschluss des freien Zyklus
                        -  B#16#04: Abschluss des Kaltstarts
                        -  B#16#05: Erster OB 1-Zyklus der neuen Master-CPU nach 
                                    Master-Reserve-Umschaltung und STOP des 
                                    bisherigen Masters *)

   #ERR := RD_SINFO (TOP_SI => #TOP_SI, START_UP_SI => #START_UP_SI);

   (* reset last_time on system startup *)
   IF #TOP_SI.EV_NUM = 1 OR #TOP_SI.EV_NUM = 2 OR #TOP_SI.EV_NUM = 4 THEN 
       #init := FALSE;
   END_IF;

   #tx := "T_PLC_MS"();
   IF #"E" AND #init THEN
       (* we need to set tl = tx when direction changes *)
       IF #DIR XOR #last_dir THEN
        #tl := #tx;
        #last_dir := #DIR;
       END_IF;
       (* check_elapsed time and calculate only if necessary *)
       IF #TR > t#0s THEN
           #"step" := DWORD_TO_DINT(SHL(IN:=DINT_TO_DWORD(DWORD_TO_DINT(#tx)-DWORD_TO_DINT(#tl)), N:=16)) / T_CONV(#TR);
       ELSE
           #"step" := 65535;
       END_IF;
       IF #"step" > 0 THEN
           (* perform the step on the ramp *)
           #tl := #tx;
           (* calculate the step response *)
           IF NOT #DIR THEN #"step" := - #"step"; END_IF;
           #RMP := DINT_TO_WORD(LIMIT(MN:=0, IN:=WORD_TO_DINT(#RMP) + #"step", MX:=65535));
       END_IF;
   ELSE
       #tl := #tx;
       #init := TRUE;
   END_IF;


   (* revison history
   hm  22. oct. 2008   rev 1.0
       original version

   hm  20. nov. 2008   rev 1.1
       set default for E to be TRUE
       added init

   *)
END_FUNCTION_BLOCK

FUNCTION_BLOCK "RMP_W"   // FB105, SCL
TITLE = RMP_W
{ S7_Optimized_Access := 'FALSE' }
AUTHOR : oscat
FAMILY : SIGGEN
NAME : RMP_W
VERSION : 2.0
// this ramp generator generates a Word wide ramp with 65535 steps
// the generator has an asynchronous set and reset
// the ramp is controlled by PT which is the total ramp time for a full sweep from 0..65535
// an UD input controlls the direction Up or Down and the E input enables the ramp generation
// a busy output indicates that the ramp is running, busy false means output is stable.
// the outputs low and high will be true when the output has reached its max or min value.
// 
// uses: _RMP_W [FB94]
//       T_PLC_MS [FC64] 
//       STIME [FB64],IDB_STIME [DB64]
   VAR_INPUT
      SET : Bool;
      PT : Time;
      "E" : Bool := TRUE;
      UP : Bool := TRUE;
      RST : Bool;
   END_VAR
   VAR_OUTPUT
      out : Word;
      busy : Bool;
      high : Bool;
      low : Bool;
   END_VAR
   VAR
      rmp : "_RMP_W";
   END_VAR
BEGIN


   #rmp(DIR := #UP, E := #"E", TR := #PT, RMP := #out);

   (* set or reset operation *)
   IF #RST THEN
       #out := 0;
   ELSIF #SET THEN
       #out := 65535;
   END_IF;

   (* checks for outputs stable and reset or set busy flag *)
   #low := #out = 0;
   #high := #out = 65535;
   #busy := NOT (#low OR #high) AND #"E";


   (* revision history:

   hm 4.10.2006        rev 1.1
       added the busy output which signals that the ramp is running.

   hm 22.1.2007        rev 1.2
       deleted unused variable step

   hm  17.9.2007       rev 1.3
       replaced time() with t_plc_ms() for compatibility reasons

   hm  28. sep 2007    rev 1.4
       added outputs on and off
       busy is now disabled while en is false
       new coding for higher accuracy and performance

   hm  5. oct 2007 rev 1.5
       added statements to allow for PT to be t#0s output jumps to max or min immediately

   hm  2. dec 2007 rev 1.6
       corrected an error in calculation of step response

   hm  25. dec 2007    rev 1.7
       corrected an error while step response was too slow for fast rise times

   hm  16. oct. 2008   rev 1.8
       improved performance

   hm  18. oct. 2008   rev 1.9
       renamed inout EN to E for compatibility reasons

   hm  23. oct. 2008   rev 2.0
       new code using _RMP_W
   *)
END_FUNCTION_BLOCK

FUNCTION_BLOCK "AIN1"   // FB106, SCL
TITLE = AIN1
{ S7_Optimized_Access := 'FALSE' }
AUTHOR : oscat
FAMILY : SIGPRO
NAME : AIN1
VERSION : 1.3
// Ain1 converts signals from A/D converters or other digital sources to an internal real value.
   VAR_INPUT
      in : DWord;
      sign_bit : Int := 255;
      error_bit : Int := 255;
      error_code_EN : Bool;
      error_code : DWord;
      overflow_bit : Int := 255;
      overflow_code_en : Bool;
      overflow_code : DWord;
      Bit_0 : Int;
      Bit_N : Int := 31;
      out_min : Real;
      out_max : Real := 1.0e+1;
      code_min : DWord;
      code_max : DWord := DW#16#FFFFFFFF;
      error_output : Real;
      overflow_output : Real := 1.0e+1;
   END_VAR
   VAR_OUTPUT
      out : Real;
      sign : Bool;
      error : Bool;
      overflow : Bool;
   END_VAR
   VAR
      tB : DWord;
      _tB AT tB : Array[0..31] of Bool;
   END_VAR
BEGIN


   (* extract error bit *)
   #error := ((SHR(IN:=#in,N:=#error_bit) AND 16#0000_0001) = 1) OR (#error_code_EN AND #error_code = #in);
   IF #error THEN
       #out := #error_output;
       RETURN;
   END_IF;

   (* strip off the data input *)
   #tB := SHR(IN:=SHL(IN:=#in, N:=31 - #Bit_N), N:=31 - #Bit_N + #Bit_0);

   (* extract overflow bit *)
   #overflow := ((SHR(IN:=#in,N:=#overflow_bit) AND 16#0000_0001) = 1) OR (#overflow_code_en AND #overflow_code = #in) OR (DWORD_TO_DINT(#tB) < DWORD_TO_DINT(#code_min) OR DWORD_TO_DINT(#tB) > DWORD_TO_DINT(#code_max));
   IF #overflow THEN
       #out := #overflow_output;
       RETURN;
   END_IF;

   (* extract sign bit *)
   #sign := (SHR(IN:=#in,N:=#sign_bit) AND 16#0000_0001) = 1;

   (* convert in to out *)
   #out := (DINT_TO_REAL(DWORD_TO_DINT(#tB) - DWORD_TO_DINT(#code_min)) * (#out_max - #out_min) / DINT_TO_REAL(DWORD_TO_DINT(#code_max) - DWORD_TO_DINT(#code_min)) + #out_min);
   IF #sign THEN #out := #out * -1.0; END_IF;



   (* revision history
   hm  23. feb 2008    rev 1.0
       original version

   hm  16. mar 2008    rev 1.1
       added type conversions to avoid warnngs under codesys 30

   hm  22. apr. 2008   rev 1.2
       corrected error in formula when code_min was set
       corrected error when sign bit was used
       optimized code for better performance

   hm  10. mar. 2009   rev 1.3
       real constants updated to new systax using dot

   *)


   (*
     (* extract error bit *)
     IF error_bit < 32 THEN
       tb := SHR(IN:=in,N:=error_bit);
       error := _tb[24]; //tb.0;
     ELSE
       error := FALSE;
     END_IF;
     (* error bit can be set or input eqals error_code if enabled *)
     error := error OR (error_code_en AND error_code = in);

     (* extract overflow bit *)
     IF overflow_bit < 32 THEN
       tb := SHR(IN:=in,N:=overflow_bit);
       overflow := _tb[24];  //tb.0;
     ELSE
       overflow := FALSE;
     END_IF;

     (* extract sign bit *)
     IF sign_bit < 32 THEN
       tB := SHR(IN:=in,N:=sign_bit);
       sign := _tb[24];  //tb.0;
     ELSE
       sign := FALSE;
     END_IF;

     (* strip off the data input *)
     tb := SHR(IN:=SHL(IN:=in,N:=31 - bit_N),N:=31 - bit_N + Bit_0);


     (* check overflow data range *)
     overflow := overflow OR (DWORD_TO_DINT(tb) < DWORD_TO_DINT(code_min) OR DWORD_TO_DINT(tb) > DWORD_TO_DINT(code_max));

     IF error THEN
       out := error_output;
     ELSIF overflow THEN
       out := overflow_output;
     ELSIF sign THEN
       out := (DWORD_TO_DINT(tb) - DWORD_TO_DINT(code_min)) * (out_max - out_min) / (DWORD_TO_DINT(code_max) - DWORD_TO_DINT(code_min)) + out_min;
     ELSE
       out := (DWORD_TO_DINT(tb) - DWORD_TO_DINT(code_min)) * (out_max - out_min) / (DWORD_TO_DINT(code_max) - DWORD_TO_DINT(code_min)) + out_min;
     END_IF;

   (* revision history
   hm  23. feb 2008    rev 1.0
       original version

   hm  16. mar 2008    rev 1.1
       added type conversions to avoid warnngs under codesys 30

   hm  22. apr. 2008   rev 1.2
       corrected error in formula when code_min was set
   *)
   *)
END_FUNCTION_BLOCK

FUNCTION_BLOCK "DELAY"   // FB107, SCL
TITLE = DELAY
{ S7_Optimized_Access := 'FALSE' }
AUTHOR : hugo
FAMILY : SIGPRO
NAME : DELAY
VERSION : 1.5
// this function block delays input values by each programm cycle
// after N+1 cycles the in value has shifted to the out.
// N can be any alue from 0 .. 32
// if n = 0 the input will be present on the output without a delay.
// f N > 32 then the output will be delayed by 32 cycles.
// any high on rst will load the buffer with in.
// 
// uses: INC1 [FC53]
   VAR_INPUT
      IN : Real;
      N : Int;
      RST : Bool;
   END_VAR
   VAR_OUTPUT
      OUT : Real;
   END_VAR
   VAR
      buf : Array[0..31] of Real;
      i : Int;
      init : Bool;
      stop : Int;
   END_VAR
BEGIN


   #stop := LIMIT(MN:=0,IN:=#N,MX:=32) - 1;
   IF #RST OR NOT #init THEN
       #init := TRUE;
       FOR #i := 0 TO #stop DO #buf[#i] := #IN; END_FOR;
       #OUT := #IN;
       #i := 0;         // Muss so sein!
   ELSIF #stop < 0 THEN
       #OUT := #IN;
   ELSE
       #OUT := #buf[#i];
       #buf[#i] := #IN;
       #i := "INC1"(X:=#i, N:=#N);
   END_IF;


   (* revision history
   hm 1.10.2006        rev 1.1
       corrected error in buffer management

   hm 19.1.2007        rev 1.2
       changed reset to load the value of in instead of 0

   hm  27. oct. 2008   rev 1.3
       improved performance

   hm  23. feb.2009    rev 1.4
       corrected an index problem

   hm  23. mar. 2009   rev 1.5
       corrected non standard write to input N

